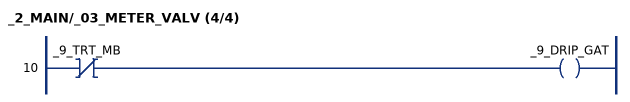
   10: XIO(_9_TRT_MB)OTE(_9_DRIP_GAT);
END_ROUTINE

ROUTINE _04_TREAT_DELY   (* ladder *)
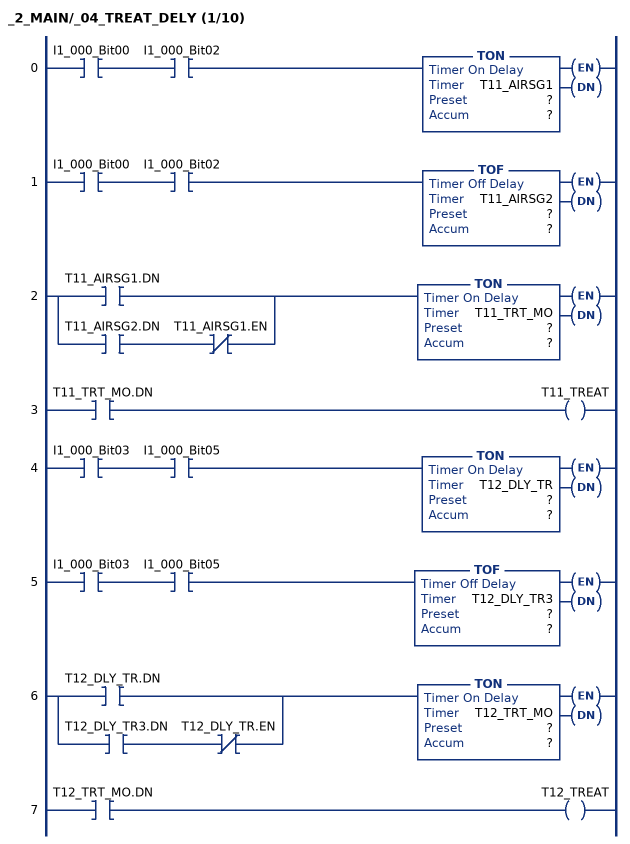
   0: XIC(I1_000_Bit00)XIC(I1_000_Bit02)TON(T11_AIRSG1,?,?);
   1: XIC(I1_000_Bit00)XIC(I1_000_Bit02)TOF(T11_AIRSG2,?,?);
   2: [XIC(T11_AIRSG1.DN) ,XIC(T11_AIRSG2.DN) XIO(T11_AIRSG1.EN) ]TON(T11_TRT_MO,?,?);
   3: XIC(T11_TRT_MO.DN)OTE(T11_TREAT);
   4: XIC(I1_000_Bit03)XIC(I1_000_Bit05)TON(T12_DLY_TR,?,?);
   5: XIC(I1_000_Bit03)XIC(I1_000_Bit05)TOF(T12_DLY_TR3,?,?);
   6: [XIC(T12_DLY_TR.DN) ,XIC(T12_DLY_TR3.DN) XIO(T12_DLY_TR.EN) ]TON(T12_TRT_MO,?,?);
   7: XIC(T12_TRT_MO.DN)OTE(T12_TREAT);
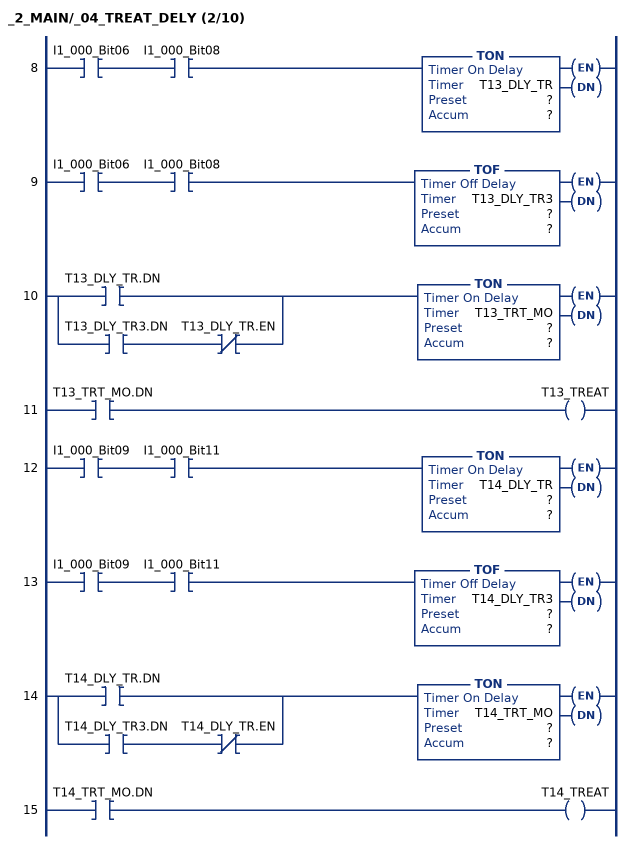
   8: XIC(I1_000_Bit06)XIC(I1_000_Bit08)TON(T13_DLY_TR,?,?);
   9: XIC(I1_000_Bit06)XIC(I1_000_Bit08)TOF(T13_DLY_TR3,?,?);
   10: [XIC(T13_DLY_TR.DN) ,XIC(T13_DLY_TR3.DN) XIO(T13_DLY_TR.EN) ]TON(T13_TRT_MO,?,?);
   11: XIC(T13_TRT_MO.DN)OTE(T13_TREAT);
   12: XIC(I1_000_Bit09)XIC(I1_000_Bit11)TON(T14_DLY_TR,?,?);
   13: XIC(I1_000_Bit09)XIC(I1_000_Bit11)TOF(T14_DLY_TR3,?,?);
   14: [XIC(T14_DLY_TR.DN) ,XIC(T14_DLY_TR3.DN) XIO(T14_DLY_TR.EN) ]TON(T14_TRT_MO,?,?);
   15: XIC(T14_TRT_MO.DN)OTE(T14_TREAT);
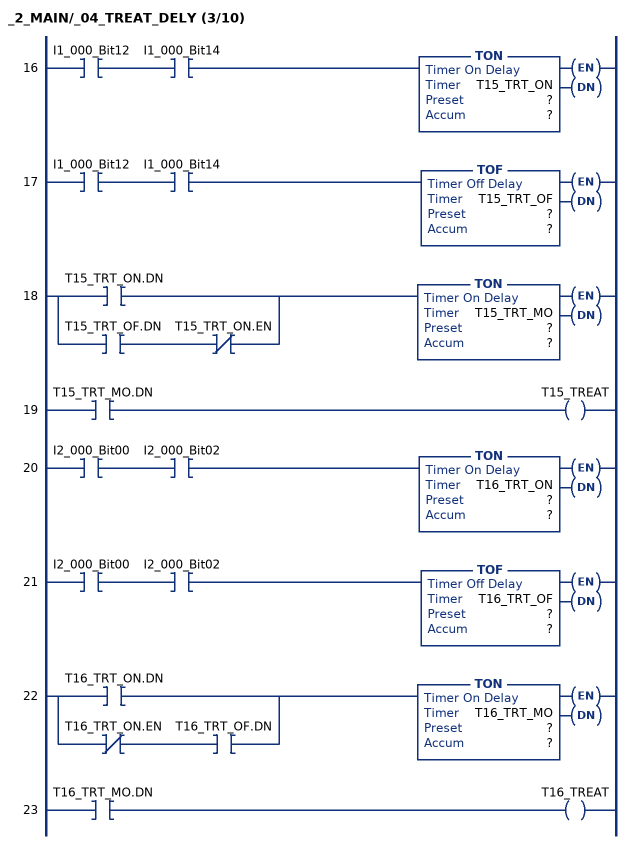
   16: XIC(I1_000_Bit12)XIC(I1_000_Bit14)TON(T15_TRT_ON,?,?);
   17: XIC(I1_000_Bit12)XIC(I1_000_Bit14)TOF(T15_TRT_OF,?,?);
   18: [XIC(T15_TRT_ON.DN) ,XIC(T15_TRT_OF.DN) XIO(T15_TRT_ON.EN) ]TON(T15_TRT_MO,?,?);
   19: XIC(T15_TRT_MO.DN)OTE(T15_TREAT);
   20: XIC(I2_000_Bit00)XIC(I2_000_Bit02)TON(T16_TRT_ON,?,?);
   21: XIC(I2_000_Bit00)XIC(I2_000_Bit02)TOF(T16_TRT_OF,?,?);
   22: [XIC(T16_TRT_ON.DN) ,XIO(T16_TRT_ON.EN) XIC(T16_TRT_OF.DN) ]TON(T16_TRT_MO,?,?);
   23: XIC(T16_TRT_MO.DN)OTE(T16_TREAT);
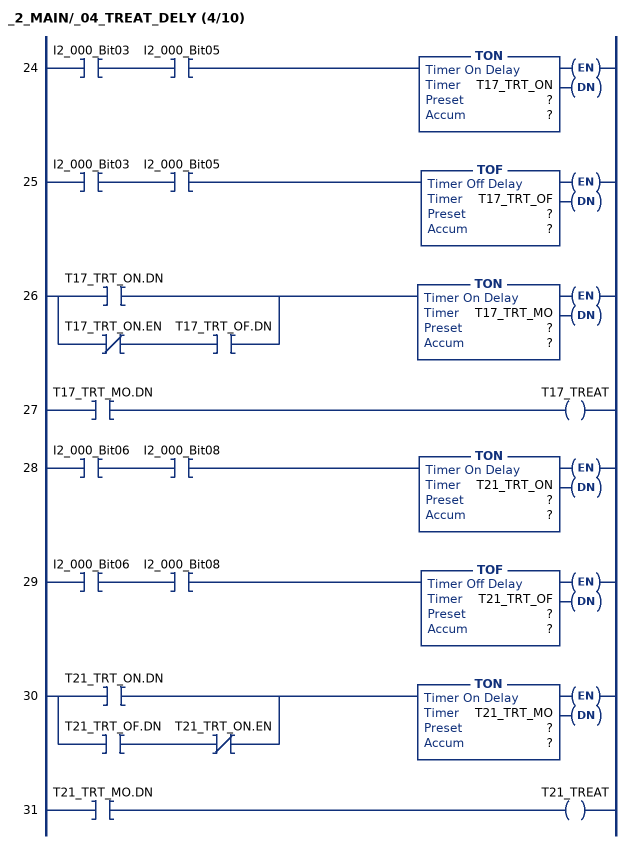
   24: XIC(I2_000_Bit03)XIC(I2_000_Bit05)TON(T17_TRT_ON,?,?);
   25: XIC(I2_000_Bit03)XIC(I2_000_Bit05)TOF(T17_TRT_OF,?,?);
   26: [XIC(T17_TRT_ON.DN) ,XIO(T17_TRT_ON.EN) XIC(T17_TRT_OF.DN) ]TON(T17_TRT_MO,?,?);
   27: XIC(T17_TRT_MO.DN)OTE(T17_TREAT);
   28: XIC(I2_000_Bit06)XIC(I2_000_Bit08)TON(T21_TRT_ON,?,?);
   29: XIC(I2_000_Bit06)XIC(I2_000_Bit08)TOF(T21_TRT_OF,?,?);
   30: [XIC(T21_TRT_ON.DN) ,XIC(T21_TRT_OF.DN) XIO(T21_TRT_ON.EN) ]TON(T21_TRT_MO,?,?);
   31: XIC(T21_TRT_MO.DN)OTE(T21_TREAT);
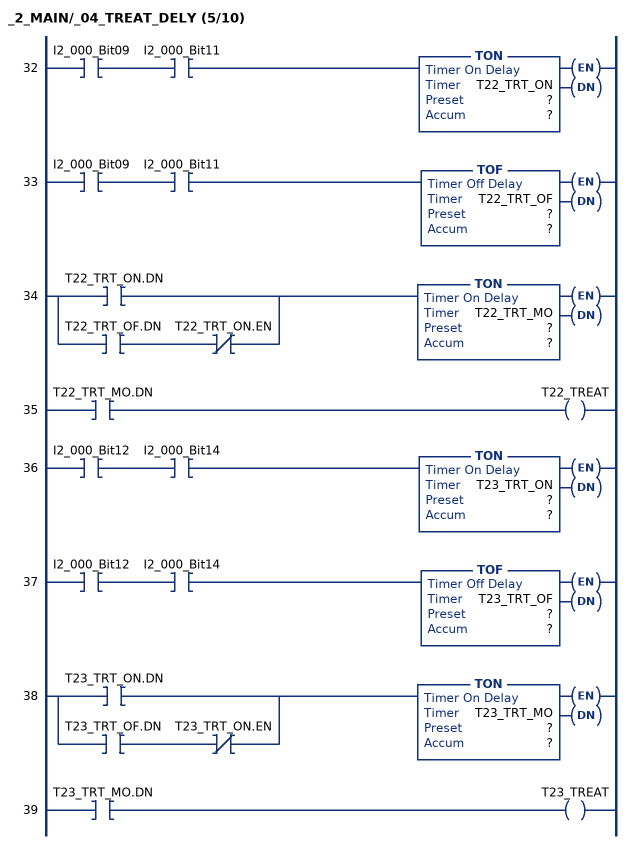
   32: XIC(I2_000_Bit09)XIC(I2_000_Bit11)TON(T22_TRT_ON,?,?);
   33: XIC(I2_000_Bit09)XIC(I2_000_Bit11)TOF(T22_TRT_OF,?,?);
   34: [XIC(T22_TRT_ON.DN) ,XIC(T22_TRT_OF.DN) XIO(T22_TRT_ON.EN) ]TON(T22_TRT_MO,?,?);
   35: XIC(T22_TRT_MO.DN)OTE(T22_TREAT);
   36: XIC(I2_000_Bit12)XIC(I2_000_Bit14)TON(T23_TRT_ON,?,?);
   37: XIC(I2_000_Bit12)XIC(I2_000_Bit14)TOF(T23_TRT_OF,?,?);
   38: [XIC(T23_TRT_ON.DN) ,XIC(T23_TRT_OF.DN) XIO(T23_TRT_ON.EN) ]TON(T23_TRT_MO,?,?);
   39: XIC(T23_TRT_MO.DN)OTE(T23_TREAT);
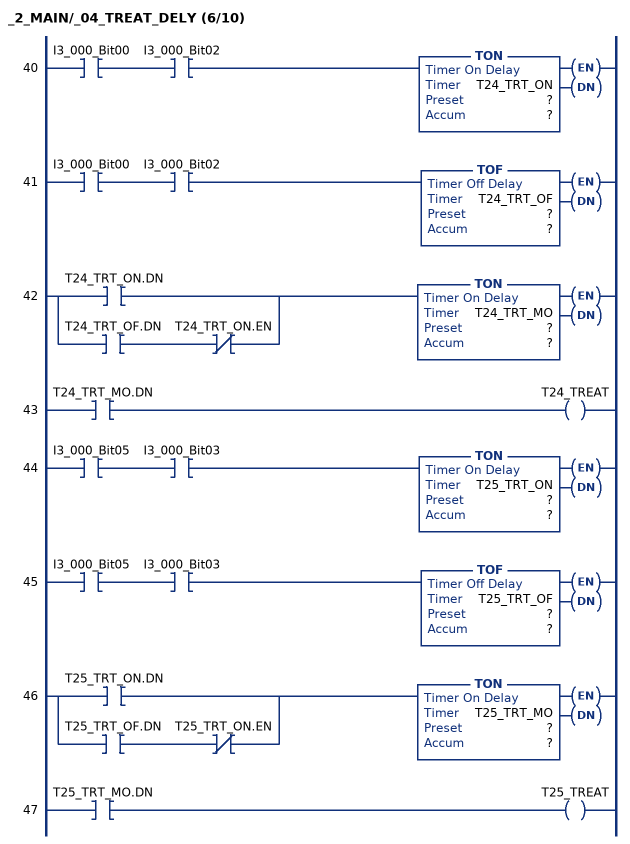
   40: XIC(I3_000_Bit00)XIC(I3_000_Bit02)TON(T24_TRT_ON,?,?);
   41: XIC(I3_000_Bit00)XIC(I3_000_Bit02)TOF(T24_TRT_OF,?,?);
   42: [XIC(T24_TRT_ON.DN) ,XIC(T24_TRT_OF.DN) XIO(T24_TRT_ON.EN) ]TON(T24_TRT_MO,?,?);
   43: XIC(T24_TRT_MO.DN)OTE(T24_TREAT);
   44: XIC(I3_000_Bit05)XIC(I3_000_Bit03)TON(T25_TRT_ON,?,?);
   45: XIC(I3_000_Bit05)XIC(I3_000_Bit03)TOF(T25_TRT_OF,?,?);
   46: [XIC(T25_TRT_ON.DN) ,XIC(T25_TRT_OF.DN) XIO(T25_TRT_ON.EN) ]TON(T25_TRT_MO,?,?);
   47: XIC(T25_TRT_MO.DN)OTE(T25_TREAT);
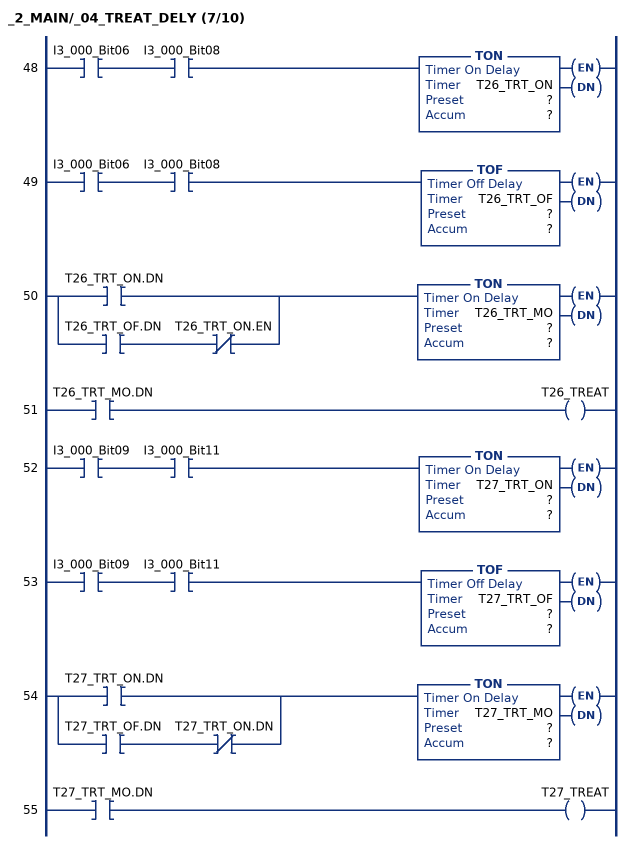
   48: XIC(I3_000_Bit06)XIC(I3_000_Bit08)TON(T26_TRT_ON,?,?);
   49: XIC(I3_000_Bit06)XIC(I3_000_Bit08)TOF(T26_TRT_OF,?,?);
   50: [XIC(T26_TRT_ON.DN) ,XIC(T26_TRT_OF.DN) XIO(T26_TRT_ON.EN) ]TON(T26_TRT_MO,?,?);
   51: XIC(T26_TRT_MO.DN)OTE(T26_TREAT);
   52: XIC(I3_000_Bit09)XIC(I3_000_Bit11)TON(T27_TRT_ON,?,?);
   53: XIC(I3_000_Bit09)XIC(I3_000_Bit11)TOF(T27_TRT_OF,?,?);
   54: [XIC(T27_TRT_ON.DN) ,XIC(T27_TRT_OF.DN) XIO(T27_TRT_ON.DN) ]TON(T27_TRT_MO,?,?);
   55: XIC(T27_TRT_MO.DN)OTE(T27_TREAT);
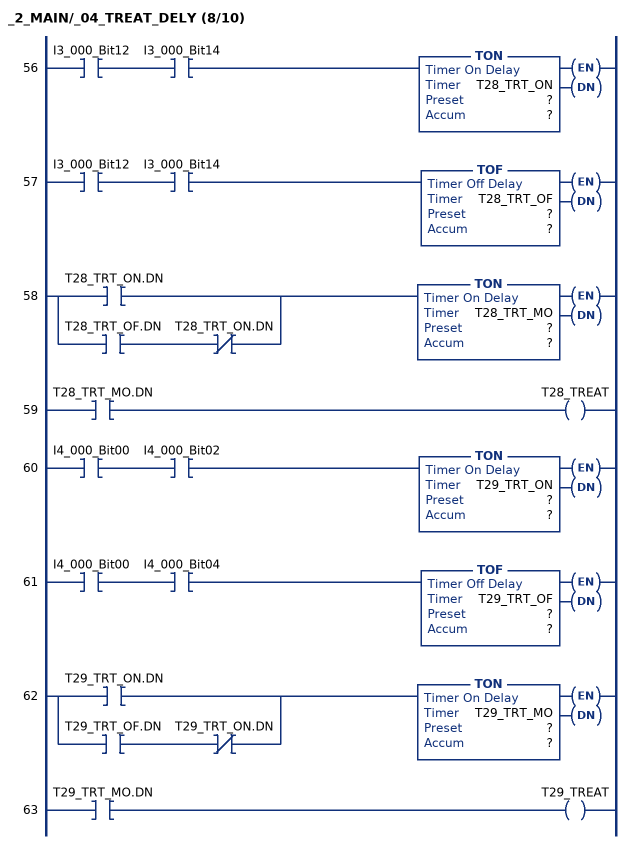
   56: XIC(I3_000_Bit12)XIC(I3_000_Bit14)TON(T28_TRT_ON,?,?);
   57: XIC(I3_000_Bit12)XIC(I3_000_Bit14)TOF(T28_TRT_OF,?,?);
   58: [XIC(T28_TRT_ON.DN) ,XIC(T28_TRT_OF.DN) XIO(T28_TRT_ON.DN) ]TON(T28_TRT_MO,?,?);
   59: XIC(T28_TRT_MO.DN)OTE(T28_TREAT);
   60: XIC(I4_000_Bit00)XIC(I4_000_Bit02)TON(T29_TRT_ON,?,?);
   61: XIC(I4_000_Bit00)XIC(I4_000_Bit04)TOF(T29_TRT_OF,?,?);
   62: [XIC(T29_TRT_ON.DN) ,XIC(T29_TRT_OF.DN) XIO(T29_TRT_ON.DN) ]TON(T29_TRT_MO,?,?);
   63: XIC(T29_TRT_MO.DN)OTE(T29_TREAT);
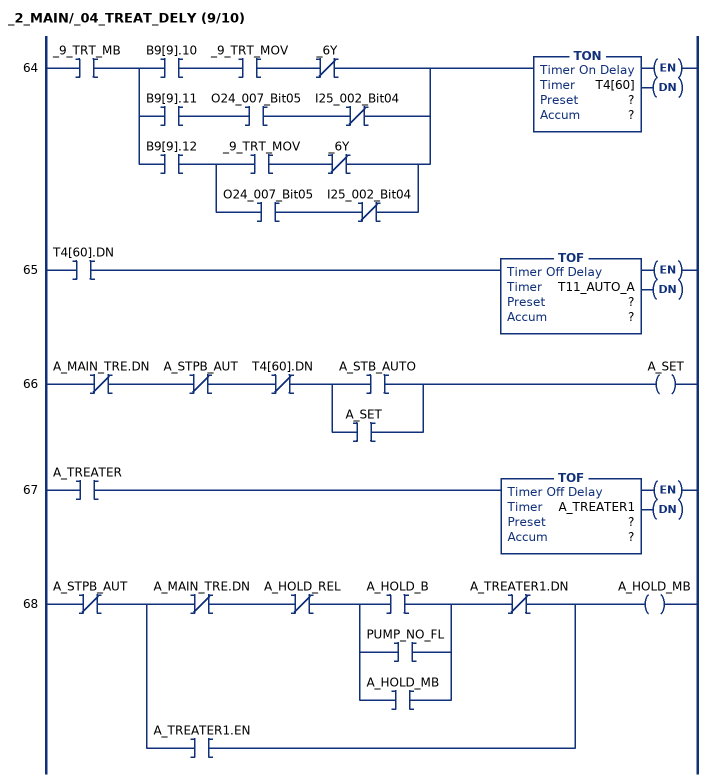
   64: XIC(_9_TRT_MB)[XIC(B9[9].10) XIC(_9_TRT_MOV) XIO(_6Y) ,XIC(B9[9].11) XIC(O24_007_Bit05) XIO(I25_002_Bit04) ,XIC(B9[9].12) [XIC(_9_TRT_MOV) XIO(_6Y) ,XIC(O24_007_Bit05) XIO(I25_002_Bit04) ] ]TON(T4[60],?,?);
   65: XIC(T4[60].DN)TOF(T11_AUTO_A,?,?);
   66: XIO(A_MAIN_TRE.DN)XIO(A_STPB_AUT)XIO(T4[60].DN)[XIC(A_STB_AUTO) ,XIC(A_SET) ]OTE(A_SET);
   67: XIC(A_TREATER)TOF(A_TREATER1,?,?);
   68: XIO(A_STPB_AUT)[XIO(A_MAIN_TRE.DN) XIO(A_HOLD_REL) [XIC(A_HOLD_B) ,XIC(PUMP_NO_FL) ,XIC(A_HOLD_MB) ] XIO(A_TREATER1.DN) ,XIC(A_TREATER1.EN) ]OTE(A_HOLD_MB);
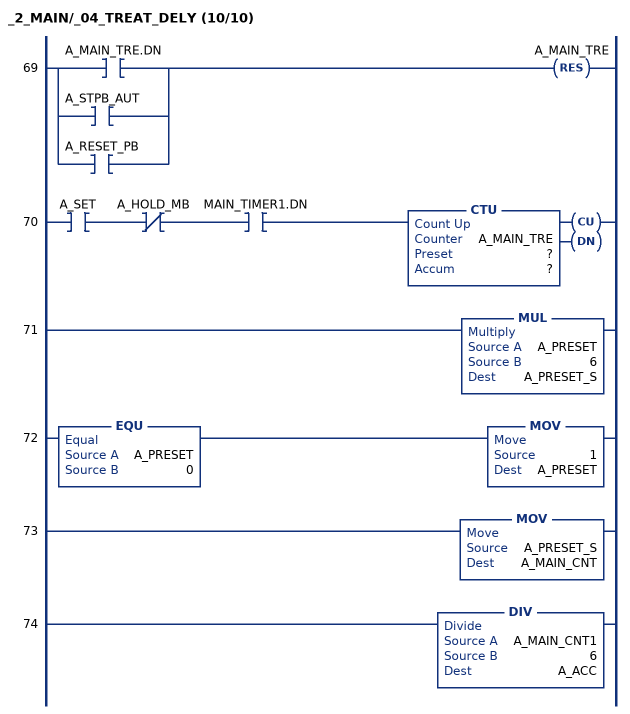
   69: [XIC(A_MAIN_TRE.DN) ,XIC(A_STPB_AUT) ,XIC(A_RESET_PB) ]RES(A_MAIN_TRE);
   70: XIC(A_SET)XIO(A_HOLD_MB)XIC(MAIN_TIMER1.DN)CTU(A_MAIN_TRE,?,?);
   71: MUL(A_PRESET,6,A_PRESET_S);
   72: EQU(A_PRESET,0)MOV(1,A_PRESET);
   73: MOV(A_PRESET_S,A_MAIN_CNT);
   74: DIV(A_MAIN_CNT1,6,A_ACC);
END_ROUTINE

ROUTINE _05_5_PMPS_ATO   (* ladder *)
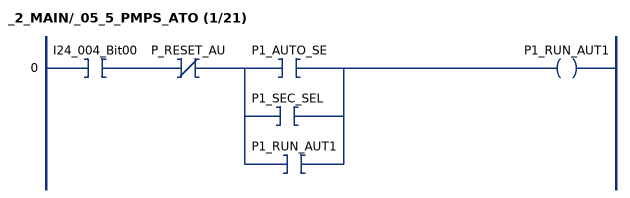
   0: XIC(I24_004_Bit00)XIO(P_RESET_AU)[XIC(P1_AUTO_SE) ,XIC(P1_SEC_SEL) ,XIC(P1_RUN_AUT1) ]OTE(P1_RUN_AUT1);
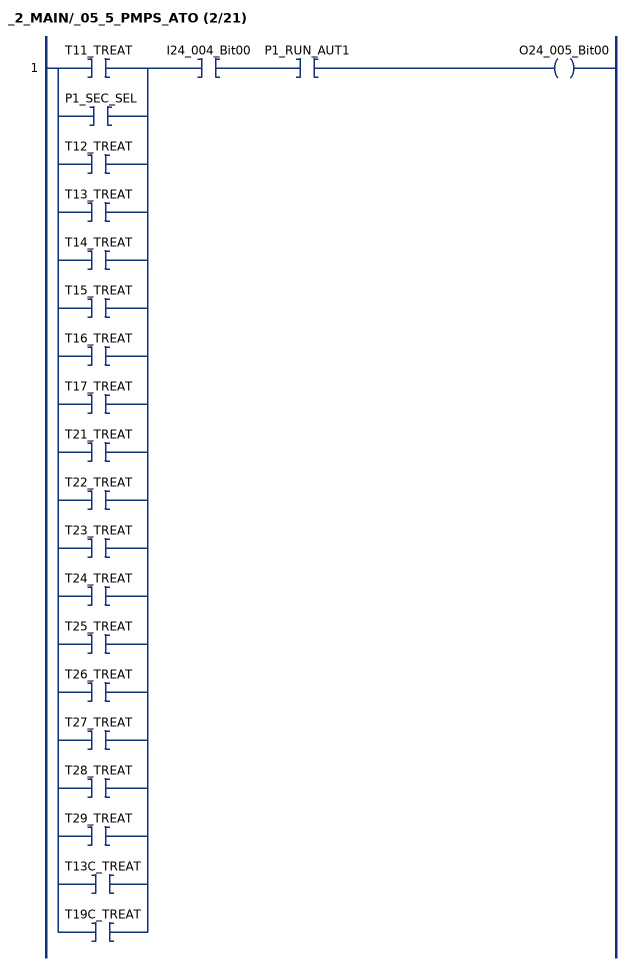
   1: [XIC(T11_TREAT) ,XIC(P1_SEC_SEL) ,XIC(T12_TREAT) ,XIC(T13_TREAT) ,XIC(T14_TREAT) ,XIC(T15_TREAT) ,XIC(T16_TREAT) ,XIC(T17_TREAT) ,XIC(T21_TREAT) ,XIC(T22_TREAT) ,XIC(T23_TREAT) ,XIC(T24_TREAT) ,XIC(T25_TREAT) ,XIC(T26_TREAT) ,XIC(T27_TREAT) ,XIC(T28_TREAT) ,XIC(T29_TREAT) ,XIC(T13C_TREAT) ,XIC(T19C_TREAT) ]XIC(I24_004_Bit00)XIC(P1_RUN_AUT1)OTE(O24_005_Bit00);
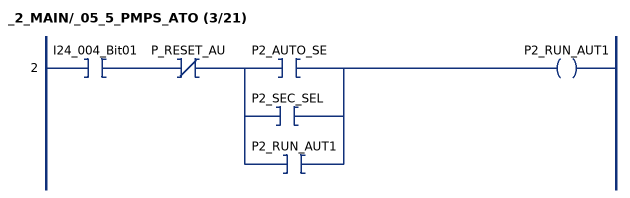
   2: XIC(I24_004_Bit01)XIO(P_RESET_AU)[XIC(P2_AUTO_SE) ,XIC(P2_SEC_SEL) ,XIC(P2_RUN_AUT1) ]OTE(P2_RUN_AUT1);
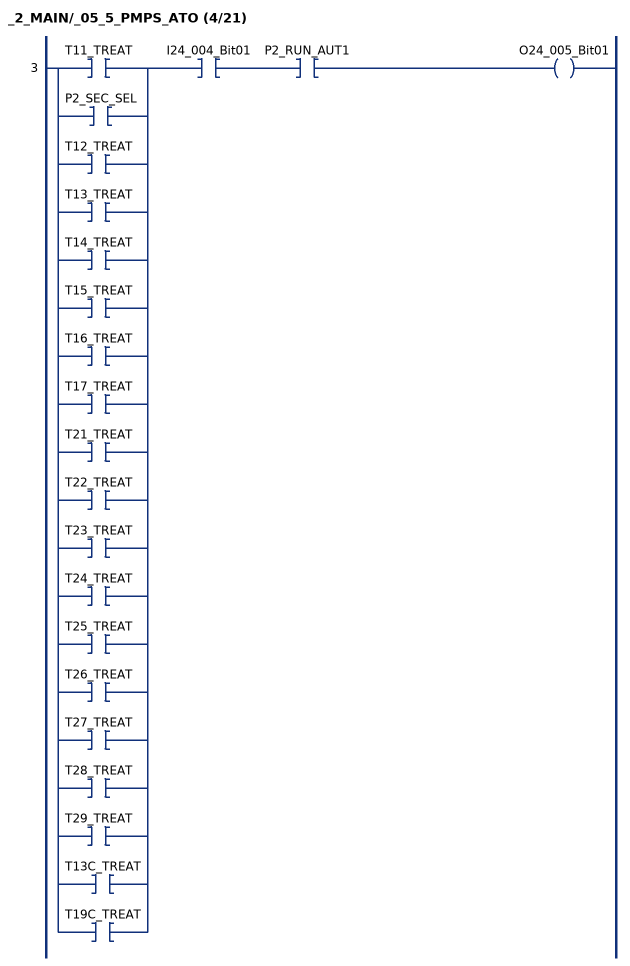
   3: [XIC(T11_TREAT) ,XIC(P2_SEC_SEL) ,XIC(T12_TREAT) ,XIC(T13_TREAT) ,XIC(T14_TREAT) ,XIC(T15_TREAT) ,XIC(T16_TREAT) ,XIC(T17_TREAT) ,XIC(T21_TREAT) ,XIC(T22_TREAT) ,XIC(T23_TREAT) ,XIC(T24_TREAT) ,XIC(T25_TREAT) ,XIC(T26_TREAT) ,XIC(T27_TREAT) ,XIC(T28_TREAT) ,XIC(T29_TREAT) ,XIC(T13C_TREAT) ,XIC(T19C_TREAT) ]XIC(I24_004_Bit01)XIC(P2_RUN_AUT1)OTE(O24_005_Bit01);
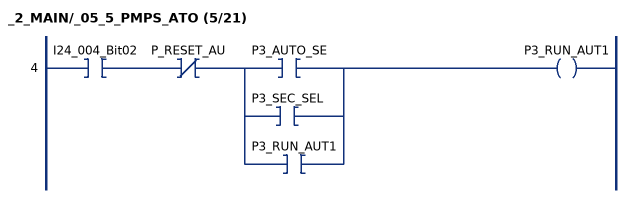
   4: XIC(I24_004_Bit02)XIO(P_RESET_AU)[XIC(P3_AUTO_SE) ,XIC(P3_SEC_SEL) ,XIC(P3_RUN_AUT1) ]OTE(P3_RUN_AUT1);
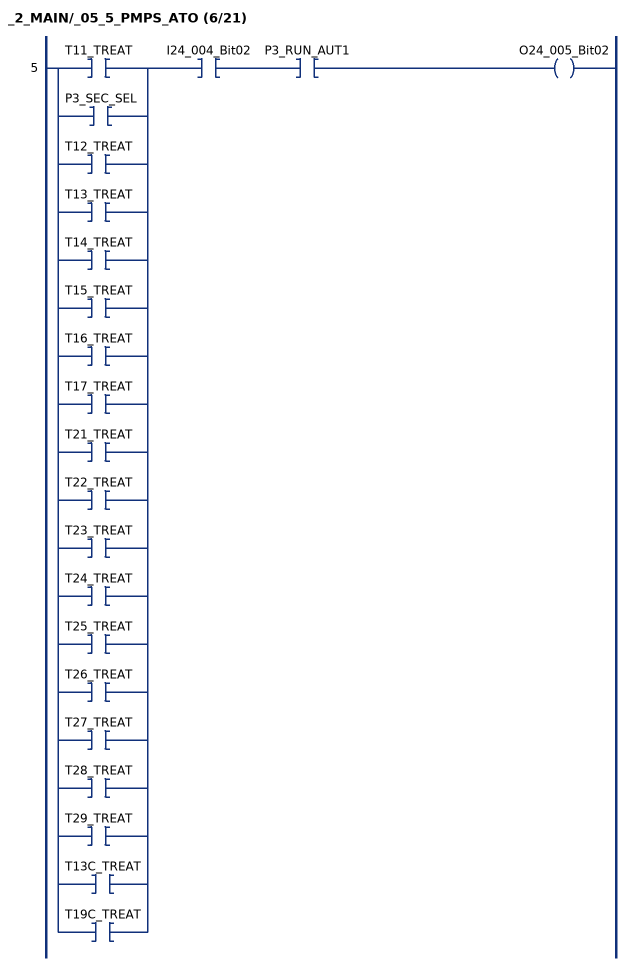
   5: [XIC(T11_TREAT) ,XIC(P3_SEC_SEL) ,XIC(T12_TREAT) ,XIC(T13_TREAT) ,XIC(T14_TREAT) ,XIC(T15_TREAT) ,XIC(T16_TREAT) ,XIC(T17_TREAT) ,XIC(T21_TREAT) ,XIC(T22_TREAT) ,XIC(T23_TREAT) ,XIC(T24_TREAT) ,XIC(T25_TREAT) ,XIC(T26_TREAT) ,XIC(T27_TREAT) ,XIC(T28_TREAT) ,XIC(T29_TREAT) ,XIC(T13C_TREAT) ,XIC(T19C_TREAT) ]XIC(I24_004_Bit02)XIC(P3_RUN_AUT1)OTE(O24_005_Bit02);
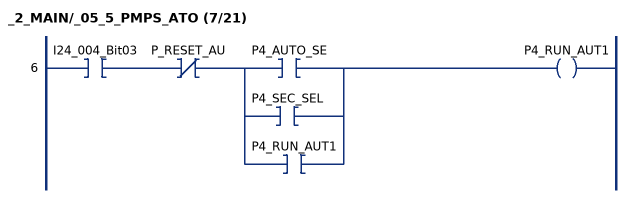
   6: XIC(I24_004_Bit03)XIO(P_RESET_AU)[XIC(P4_AUTO_SE) ,XIC(P4_SEC_SEL) ,XIC(P4_RUN_AUT1) ]OTE(P4_RUN_AUT1);
